(* Logix 5000 project; controller PLC_MCC1300_75F1 vendor 1 type 14 code 166 rev 32.11; software revision 32.04; part 26 of 83 *)
(* tags used below, declared in another part *)
   CM_LineToConveyorStacker_JS2 : CM_LineToConveyorStacker;
   GP_OB_InitializeMain : GP_OB_Initialize;
   M302SpeedUp : MAC_SpeedUp;
   M317 : MAC_Conveyor_Single;
   M317_Data : UDT_Convoy_SL;
   M317_HMW : MAC_Conveyor_HMW;
   M317_M3_ChangeSpeed : BOOL;
   M317_M3_DR_IN_MAJ : MOTION_INSTRUCTION;
   M317_M3_DR_L : AXIS_CIP_DRIVE;
   M317_M3_DR_OUT_MAJ : MOTION_INSTRUCTION;
   M317_M3_DR_OUT_MAS : MOTION_INSTRUCTION;
   M317_M3_DR_OUT_MCD : MOTION_INSTRUCTION;
   M317_SpaceConv_Utilities : SpaceConv_Utilities;
   M350Popup : MAC_Popup_ZC;
   M351 : MAC_Conveyor;
   M351_ALM : MAC_Conveyor_ALM;
   M351_Data : UDT_Convoy_SL;
   M351_HMR : MAC_Conveyor_HMR;
   M351_HMW : MAC_Conveyor_HMW;
   M351_M1_DR : AXIS_CIP_DRIVE;
   M351_M1_DR_IN_MAJ : MOTION_INSTRUCTION;
   M351_M1_DR_IN_MAR : MOTION_INSTRUCTION;
   M351_M1_DR_IN_MAS : MOTION_INSTRUCTION;
   M351_M1_DR_IN_MRP : MOTION_INSTRUCTION;
   M351_M1_DR_MAFR : MOTION_INSTRUCTION;
   M351_M1_DR_MDR : MOTION_INSTRUCTION;
   M351_M1_DR_MSF : MOTION_INSTRUCTION;
   M351_M1_DR_MSO : MOTION_INSTRUCTION;
   M351_M1_DR_OUT_MAJ : MOTION_INSTRUCTION;
   M351_M1_DR_OUT_MAM : MOTION_INSTRUCTION;
   M351_M1_DR_OUT_MAR : MOTION_INSTRUCTION;
   M351_M1_DR_OUT_MAS : MOTION_INSTRUCTION;
   M351_M1_DR_OUT_MCD : MOTION_INSTRUCTION;
   M351_M1_DR_OUT_MRP : MOTION_INSTRUCTION;
   M351_SpaceConv_Utilities : SpaceConv_Utilities;
   M352 : MAC_Conveyor;
   TMP_d : DINT;
   TMP_dDirection : DINT;
   TMP_r : REAL;
   TMP_rAcc : REAL;
   TMP_rDec : REAL;
   TMP_rSpeed : REAL;
   TMP_rTarget_M2 : REAL;
   TMP_xForwardCommadnForCleaningZone : BOOL;
   TMP_xPositioning : BOOL;
   TMP_xPositioning_M2 : BOOL;
   TMP_xPositioning_M3 : BOOL;
   TMP_xPowerSaving : BOOL;
   TMP_xReverse : BOOL;
   TMP_xReverse_M2 : BOOL;
   TMP_xReverse_M3 : BOOL;
   TMP_xRun : BOOL;
   TMP_xRun_M2 : BOOL;
   TMP_xRun_M3 : BOOL;
   xAlwaysOFF : BOOL;
   xDebugOFF : BOOL;
   Z300_Conveyor : UDT_StandConv[29];
   Z300_Conveyor_Conf : UDT_Conveyor_Config[29];
   Z300_Conveyor_HMW : MAC_Conveyor_ZC_HMW[29];
   Z300_Conveyor_IN_MOTION : MAC_Conveyor_ZC_IN_MOTION[29];
   Z301_HMR : MAC_Zone_ML_HMR;
   Z402 : MAC_Zone;
   Z900 : MAC_Zone;
   Z900_HMW : MAC_Zone_HMW;
(* CommandLogic, continued *)

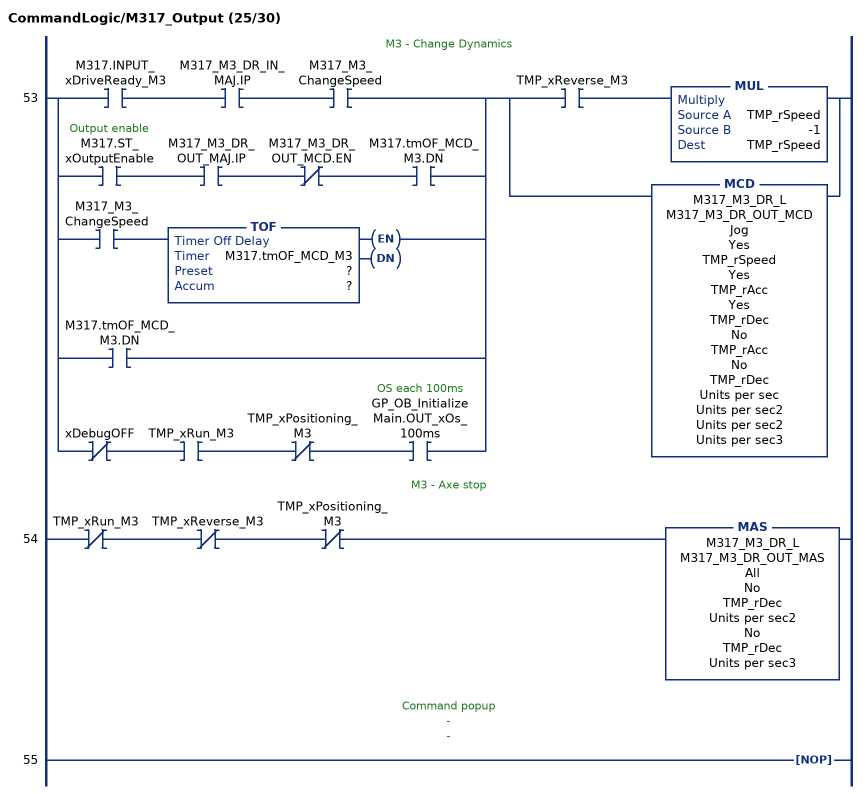
   [picture p307: CommandLogic/M317_Output rungs 53-55]
   // M3 - Change Dynamics
   53: [XIC(M317.INPUT_xDriveReady_M3) XIC(M317_M3_DR_IN_MAJ.IP) XIC(M317_M3_ChangeSpeed) ,XIC(M317.ST_xOutputEnable) XIC(M317_M3_DR_OUT_MAJ.IP) XIO(M317_M3_DR_OUT_MCD.EN) XIC(M317.tmOF_MCD_M3.DN) ,[XIC(M317_M3_ChangeSpeed) TOF(M317.tmOF_MCD_M3,?,?) ,XIC(M317.tmOF_MCD_M3.DN) ] ,XIO(xDebugOFF) XIC(TMP_xRun_M3) XIO(TMP_xPositioning_M3) XIC(GP_OB_InitializeMain.OUT_xOs_100ms) ][XIC(TMP_xReverse_M3) MUL(TMP_rSpeed,-1,TMP_rSpeed) ,MCD(M317_M3_DR_L,M317_M3_DR_OUT_MCD,Jog,Yes,TMP_rSpeed,Yes,TMP_rAcc,Yes,TMP_rDec,No,TMP_rAcc,No,TMP_rDec,Units per sec,Units per sec2,Units per sec2,Units per sec3) ];
   // M3 - Axe stop
   54: XIO(TMP_xRun_M3)XIO(TMP_xReverse_M3)XIO(TMP_xPositioning_M3)MAS(M317_M3_DR_L,M317_M3_DR_OUT_MAS,All,No,TMP_rDec,Units per sec2,No,TMP_rDec,Units per sec3);
   // Command popup
   // -
   // -
   55: NOP();
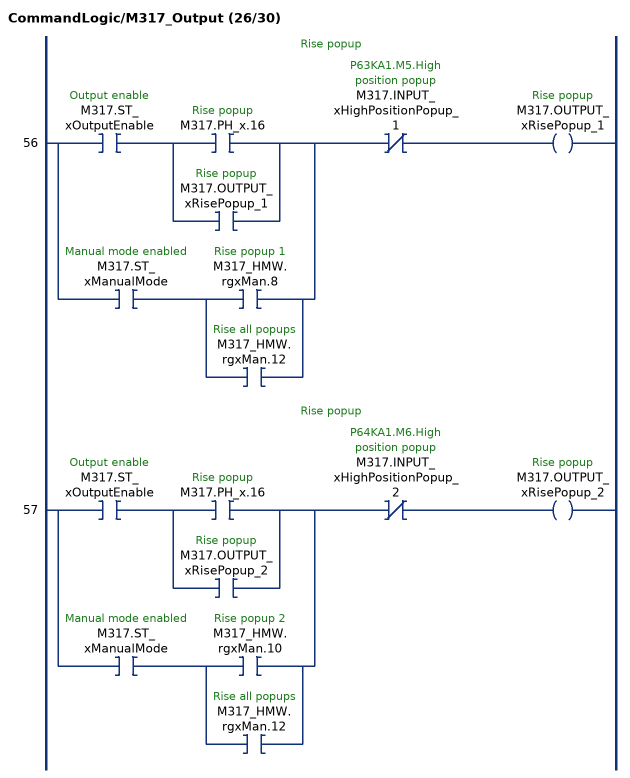
   // Rise popup
   56: [XIC(M317.ST_xOutputEnable) [XIC(M317.PH_x.16) ,XIC(M317.OUTPUT_xRisePopup_1) ] ,XIC(M317.ST_xManualMode) [XIC(M317_HMW.rgxMan.8) ,XIC(M317_HMW.rgxMan.12) ] ]XIO(M317.INPUT_xHighPositionPopup_1)OTE(M317.OUTPUT_xRisePopup_1);
   // Rise popup
   57: [XIC(M317.ST_xOutputEnable) [XIC(M317.PH_x.16) ,XIC(M317.OUTPUT_xRisePopup_2) ] ,XIC(M317.ST_xManualMode) [XIC(M317_HMW.rgxMan.10) ,XIC(M317_HMW.rgxMan.12) ] ]XIO(M317.INPUT_xHighPositionPopup_2)OTE(M317.OUTPUT_xRisePopup_2);
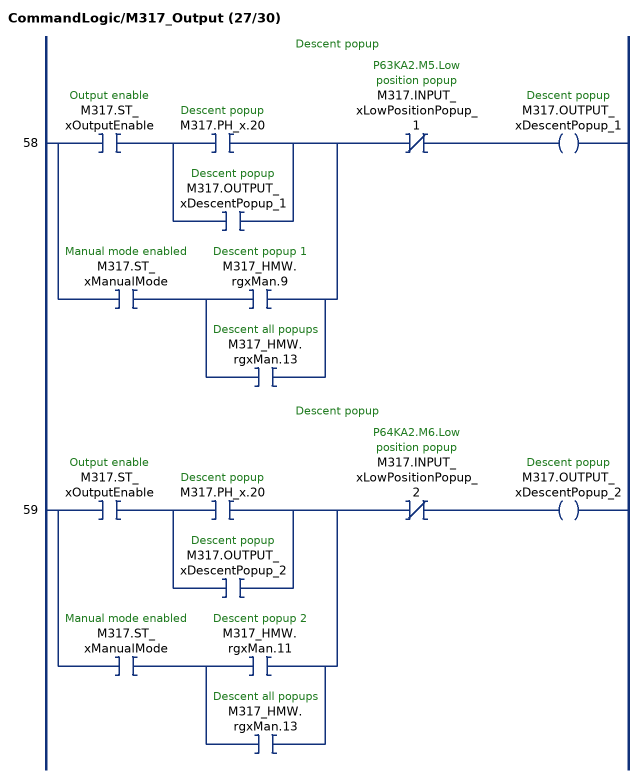
   // Descent popup
   58: [XIC(M317.ST_xOutputEnable) [XIC(M317.PH_x.20) ,XIC(M317.OUTPUT_xDescentPopup_1) ] ,XIC(M317.ST_xManualMode) [XIC(M317_HMW.rgxMan.9) ,XIC(M317_HMW.rgxMan.13) ] ]XIO(M317.INPUT_xLowPositionPopup_1)OTE(M317.OUTPUT_xDescentPopup_1);
   // Descent popup
   59: [XIC(M317.ST_xOutputEnable) [XIC(M317.PH_x.20) ,XIC(M317.OUTPUT_xDescentPopup_2) ] ,XIC(M317.ST_xManualMode) [XIC(M317_HMW.rgxMan.11) ,XIC(M317_HMW.rgxMan.13) ] ]XIO(M317.INPUT_xLowPositionPopup_2)OTE(M317.OUTPUT_xDescentPopup_2);
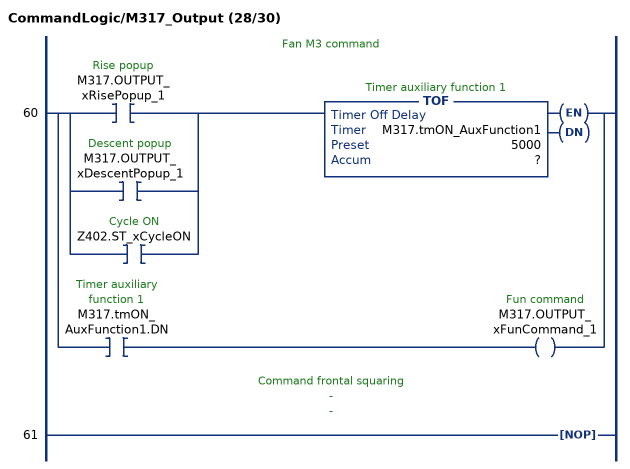
   // Fan M3 command
   60: [[XIC(M317.OUTPUT_xRisePopup_1) ,[XIC(M317.OUTPUT_xDescentPopup_1) ,XIC(Z402.ST_xCycleON) ] ] TOF(M317.tmON_AuxFunction1,?,?) ,XIC(M317.tmON_AuxFunction1.DN) OTE(M317.OUTPUT_xFunCommand_1) ];
   // Command frontal squaring
   // -
   // -
   61: NOP();
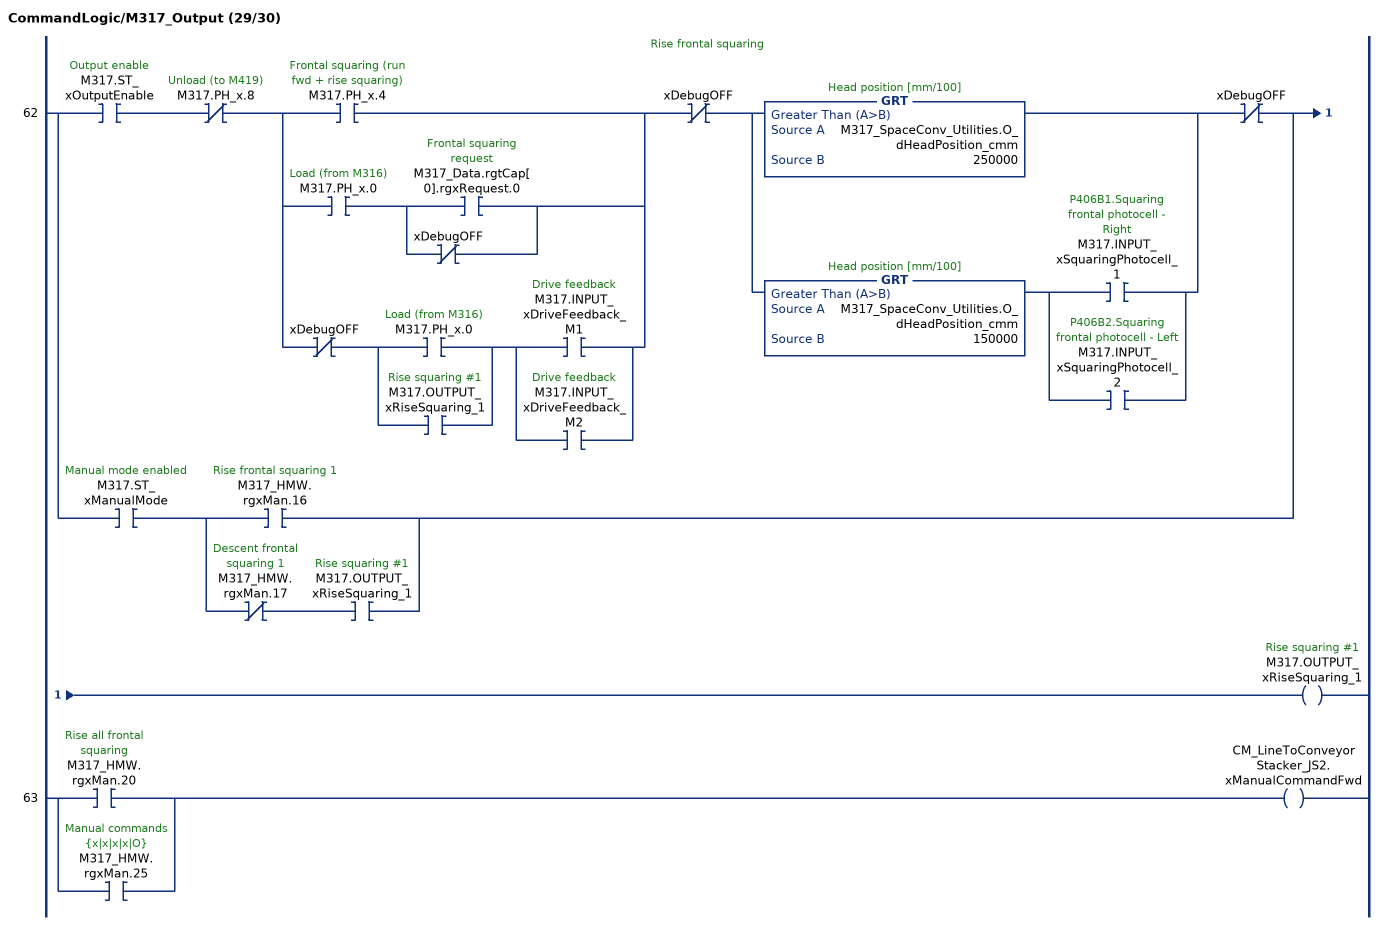
   // Rise frontal squaring
   62: [XIC(M317.ST_xOutputEnable) XIO(M317.PH_x.8) [XIC(M317.PH_x.4) ,XIC(M317.PH_x.0) [XIC(M317_Data.rgtCap[0].rgxRequest.0) ,XIO(xDebugOFF) ] ,XIO(xDebugOFF) [XIC(M317.PH_x.0) ,XIC(M317.OUTPUT_xRiseSquaring_1) ] [XIC(M317.INPUT_xDriveFeedback_M1) ,XIC(M317.INPUT_xDriveFeedback_M2) ] ] XIO(xDebugOFF) [GRT(M317_SpaceConv_Utilities.O_dHeadPosition_cmm,250000) ,GRT(M317_SpaceConv_Utilities.O_dHeadPosition_cmm,150000) [XIC(M317.INPUT_xSquaringPhotocell_1) ,XIC(M317.INPUT_xSquaringPhotocell_2) ] ] XIO(xDebugOFF) ,XIC(M317.ST_xManualMode) [XIC(M317_HMW.rgxMan.16) ,XIO(M317_HMW.rgxMan.17) XIC(M317.OUTPUT_xRiseSquaring_1) ] ]OTE(M317.OUTPUT_xRiseSquaring_1);
   63: [XIC(M317_HMW.rgxMan.20) ,XIC(M317_HMW.rgxMan.25) ]OTE(CM_LineToConveyorStacker_JS2.xManualCommandFwd);
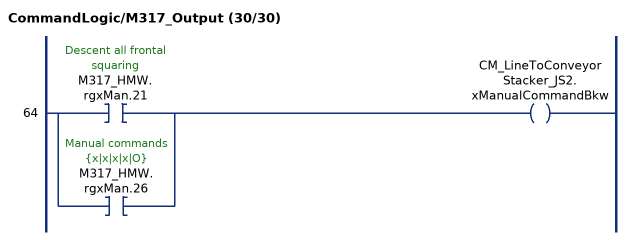
   64: [XIC(M317_HMW.rgxMan.21) ,XIC(M317_HMW.rgxMan.26) ]OTE(CM_LineToConveyorStacker_JS2.xManualCommandBkw);
END_ROUTINE

ROUTINE M350M1_Conveyor_Output   (* ladder *)
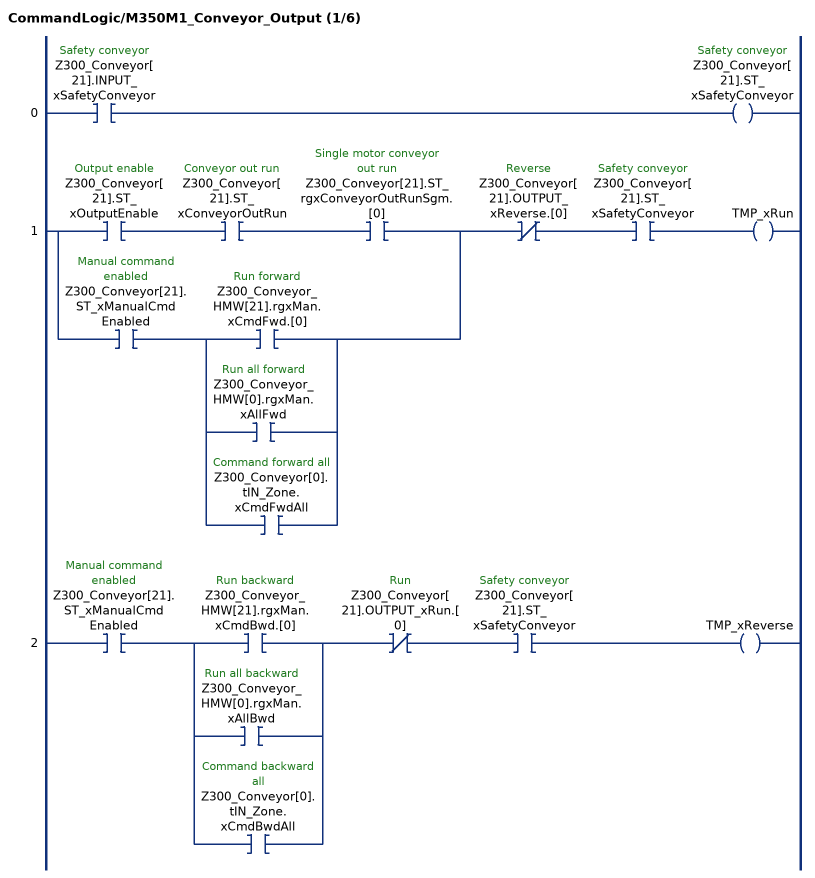
   0: XIC(Z300_Conveyor[21].INPUT_xSafetyConveyor)OTE(Z300_Conveyor[21].ST_xSafetyConveyor);
   1: [XIC(Z300_Conveyor[21].ST_xOutputEnable) XIC(Z300_Conveyor[21].ST_xConveyorOutRun) XIC(Z300_Conveyor[21].ST_rgxConveyorOutRunSgm.[0]) ,XIC(Z300_Conveyor[21].ST_xManualCmdEnabled) [XIC(Z300_Conveyor_HMW[21].rgxMan.xCmdFwd.[0]) ,XIC(Z300_Conveyor_HMW[0].rgxMan.xAllFwd) ,XIC(Z300_Conveyor[0].tIN_Zone.xCmdFwdAll) ] ]XIO(Z300_Conveyor[21].OUTPUT_xReverse.[0])XIC(Z300_Conveyor[21].ST_xSafetyConveyor)OTE(TMP_xRun);
   2: XIC(Z300_Conveyor[21].ST_xManualCmdEnabled)[XIC(Z300_Conveyor_HMW[21].rgxMan.xCmdBwd.[0]) ,XIC(Z300_Conveyor_HMW[0].rgxMan.xAllBwd) ,XIC(Z300_Conveyor[0].tIN_Zone.xCmdBwdAll) ]XIO(Z300_Conveyor[21].OUTPUT_xRun.[0])XIC(Z300_Conveyor[21].ST_xSafetyConveyor)OTE(TMP_xReverse);
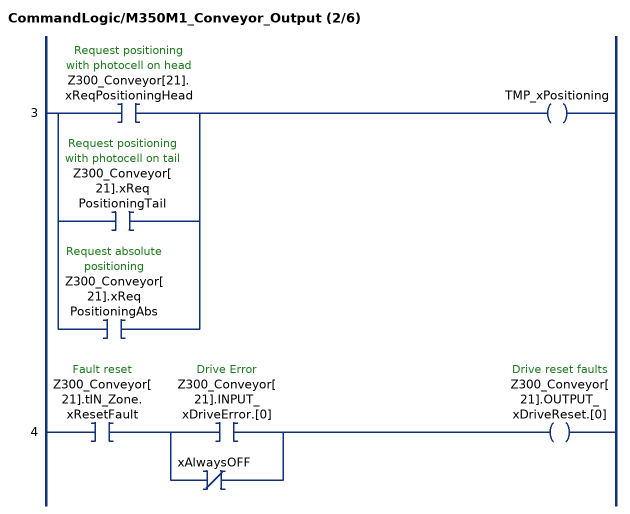
   3: [XIC(Z300_Conveyor[21].xReqPositioningHead) ,XIC(Z300_Conveyor[21].xReqPositioningTail) ,XIC(Z300_Conveyor[21].xReqPositioningAbs) ]OTE(TMP_xPositioning);
   4: XIC(Z300_Conveyor[21].tIN_Zone.xResetFault)[XIC(Z300_Conveyor[21].INPUT_xDriveError.[0]) ,XIO(xAlwaysOFF) ]OTE(Z300_Conveyor[21].OUTPUT_xDriveReset.[0]);
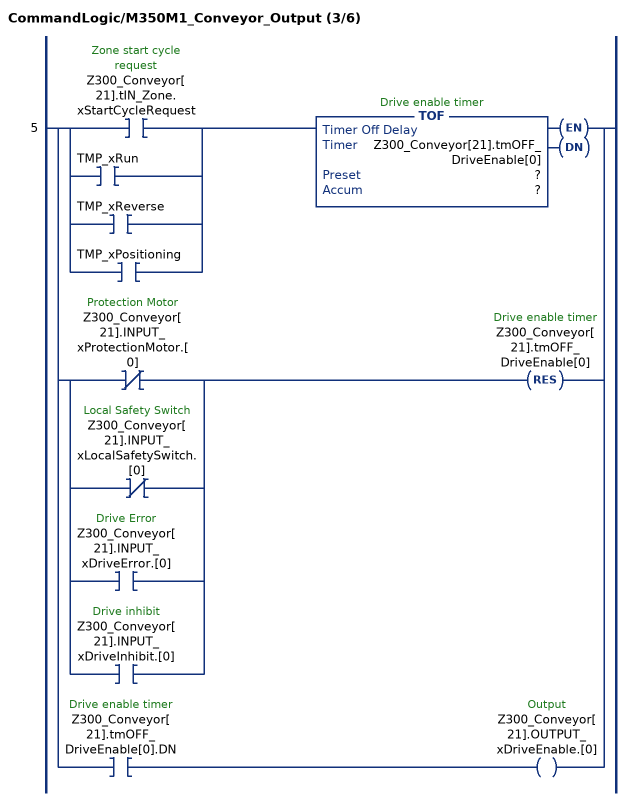
   5: [[XIC(Z300_Conveyor[21].tIN_Zone.xStartCycleRequest) ,XIC(TMP_xRun) ,XIC(TMP_xReverse) ,XIC(TMP_xPositioning) ] TOF(Z300_Conveyor[21].tmOFF_DriveEnable[0],?,?) ,[XIO(Z300_Conveyor[21].INPUT_xProtectionMotor.[0]) ,XIO(Z300_Conveyor[21].INPUT_xLocalSafetySwitch.[0]) ,XIC(Z300_Conveyor[21].INPUT_xDriveError.[0]) ,XIC(Z300_Conveyor[21].INPUT_xDriveInhibit.[0]) ] RES(Z300_Conveyor[21].tmOFF_DriveEnable[0]) ,XIC(Z300_Conveyor[21].tmOFF_DriveEnable[0].DN) OTE(Z300_Conveyor[21].OUTPUT_xDriveEnable.[0]) ];
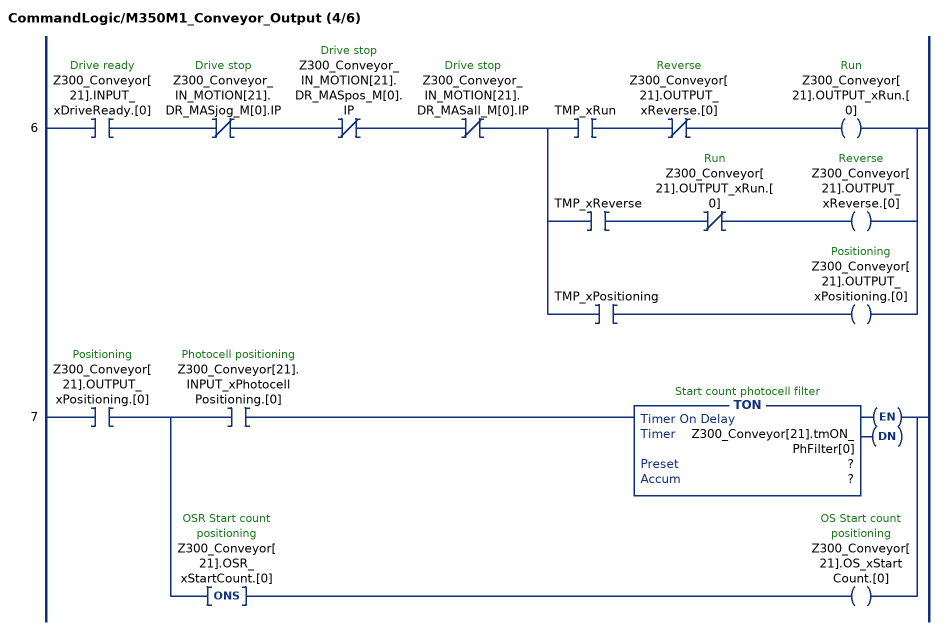
   6: XIC(Z300_Conveyor[21].INPUT_xDriveReady.[0])XIO(Z300_Conveyor_IN_MOTION[21].DR_MASjog_M[0].IP)XIO(Z300_Conveyor_IN_MOTION[21].DR_MASpos_M[0].IP)XIO(Z300_Conveyor_IN_MOTION[21].DR_MASall_M[0].IP)[XIC(TMP_xRun) XIO(Z300_Conveyor[21].OUTPUT_xReverse.[0]) OTE(Z300_Conveyor[21].OUTPUT_xRun.[0]) ,XIC(TMP_xReverse) XIO(Z300_Conveyor[21].OUTPUT_xRun.[0]) OTE(Z300_Conveyor[21].OUTPUT_xReverse.[0]) ,XIC(TMP_xPositioning) OTE(Z300_Conveyor[21].OUTPUT_xPositioning.[0]) ];
   7: XIC(Z300_Conveyor[21].OUTPUT_xPositioning.[0])[XIC(Z300_Conveyor[21].INPUT_xPhotocellPositioning.[0]) TON(Z300_Conveyor[21].tmON_PhFilter[0],?,?) ,ONS(Z300_Conveyor[21].OSR_xStartCount.[0]) OTE(Z300_Conveyor[21].OS_xStartCount.[0]) ];
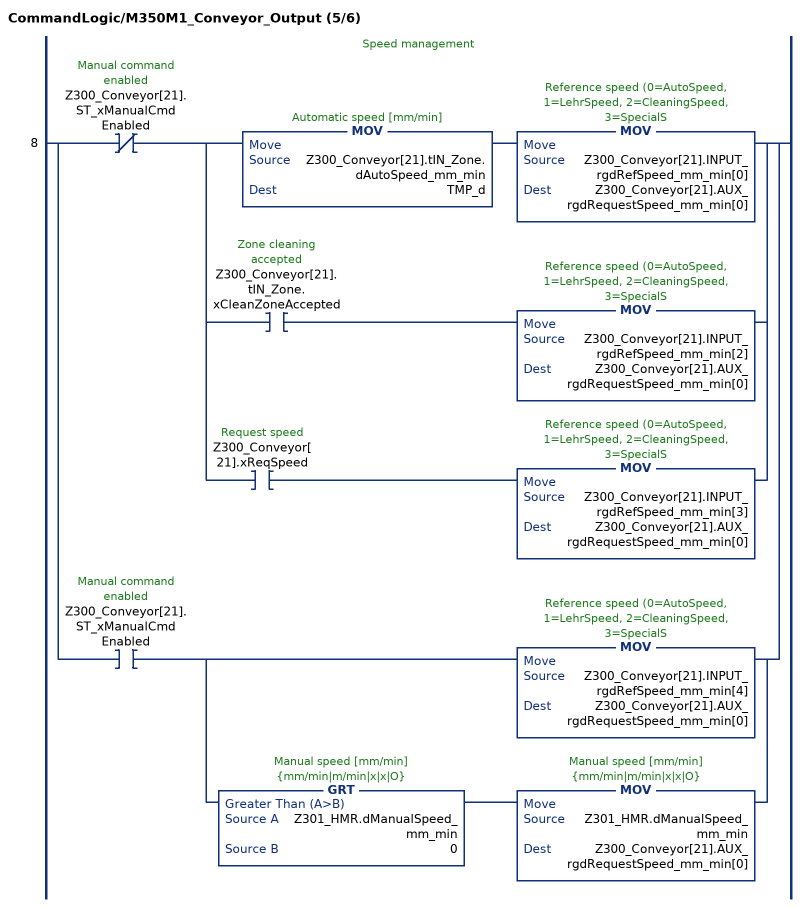
   // Speed management
   8: [XIO(Z300_Conveyor[21].ST_xManualCmdEnabled) [MOV(Z300_Conveyor[21].tIN_Zone.dAutoSpeed_mm_min,TMP_d) MOV(Z300_Conveyor[21].INPUT_rgdRefSpeed_mm_min[0],Z300_Conveyor[21].AUX_rgdRequestSpeed_mm_min[0]) ,XIC(Z300_Conveyor[21].tIN_Zone.xCleanZoneAccepted) MOV(Z300_Conveyor[21].INPUT_rgdRefSpeed_mm_min[2],Z300_Conveyor[21].AUX_rgdRequestSpeed_mm_min[0]) ,XIC(Z300_Conveyor[21].xReqSpeed) MOV(Z300_Conveyor[21].INPUT_rgdRefSpeed_mm_min[3],Z300_Conveyor[21].AUX_rgdRequestSpeed_mm_min[0]) ] ,XIC(Z300_Conveyor[21].ST_xManualCmdEnabled) [MOV(Z300_Conveyor[21].INPUT_rgdRefSpeed_mm_min[4],Z300_Conveyor[21].AUX_rgdRequestSpeed_mm_min[0]) ,GRT(Z301_HMR.dManualSpeed_mm_min,0) MOV(Z301_HMR.dManualSpeed_mm_min,Z300_Conveyor[21].AUX_rgdRequestSpeed_mm_min[0]) ] ];
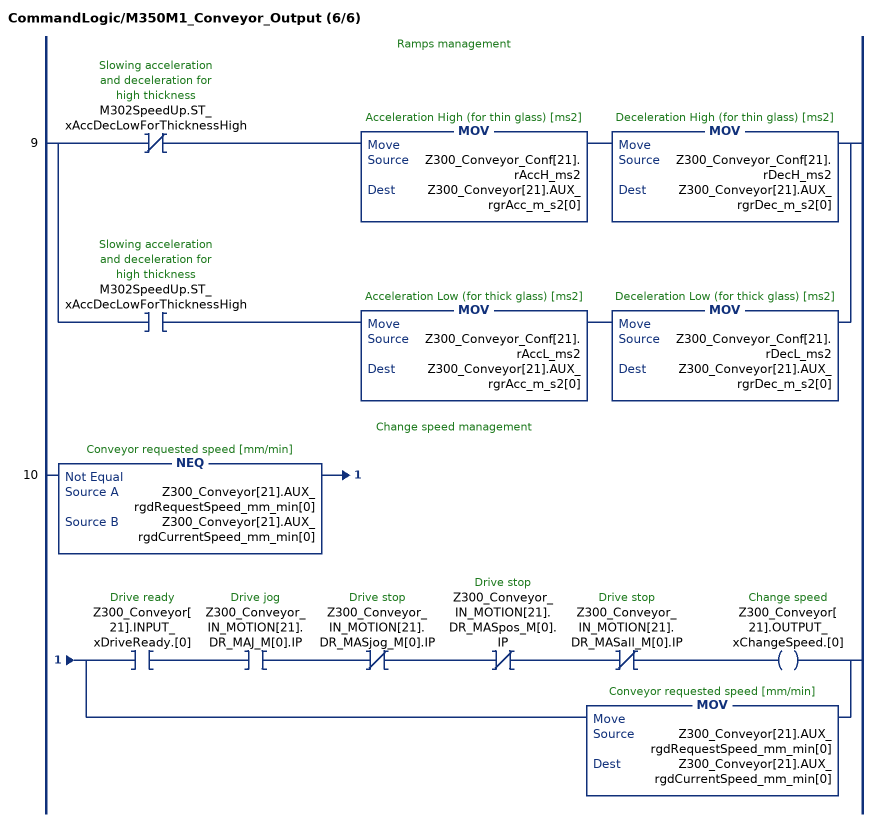
   // Ramps management
   9: [XIO(M302SpeedUp.ST_xAccDecLowForThicknessHigh) MOV(Z300_Conveyor_Conf[21].rAccH_ms2,Z300_Conveyor[21].AUX_rgrAcc_m_s2[0]) MOV(Z300_Conveyor_Conf[21].rDecH_ms2,Z300_Conveyor[21].AUX_rgrDec_m_s2[0]) ,XIC(M302SpeedUp.ST_xAccDecLowForThicknessHigh) MOV(Z300_Conveyor_Conf[21].rAccL_ms2,Z300_Conveyor[21].AUX_rgrAcc_m_s2[0]) MOV(Z300_Conveyor_Conf[21].rDecL_ms2,Z300_Conveyor[21].AUX_rgrDec_m_s2[0]) ];
   // Change speed management
   10: NEQ(Z300_Conveyor[21].AUX_rgdRequestSpeed_mm_min[0],Z300_Conveyor[21].AUX_rgdCurrentSpeed_mm_min[0])[XIC(Z300_Conveyor[21].INPUT_xDriveReady.[0]) XIC(Z300_Conveyor_IN_MOTION[21].DR_MAJ_M[0].IP) XIO(Z300_Conveyor_IN_MOTION[21].DR_MASjog_M[0].IP) XIO(Z300_Conveyor_IN_MOTION[21].DR_MASpos_M[0].IP) XIO(Z300_Conveyor_IN_MOTION[21].DR_MASall_M[0].IP) OTE(Z300_Conveyor[21].OUTPUT_xChangeSpeed.[0]) ,MOV(Z300_Conveyor[21].AUX_rgdRequestSpeed_mm_min[0],Z300_Conveyor[21].AUX_rgdCurrentSpeed_mm_min[0]) ];
END_ROUTINE

ROUTINE M351_Output   (* ladder *)
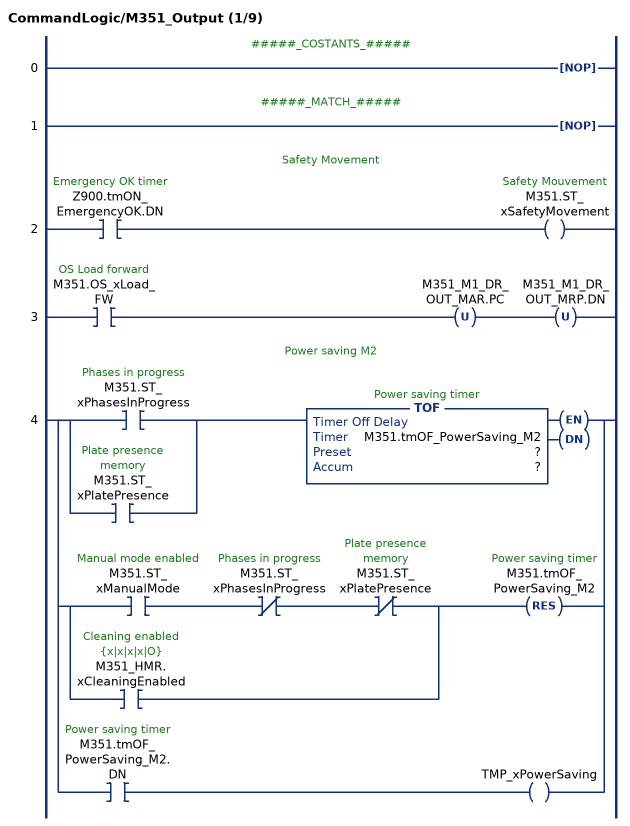
   // #####_COSTANTS_#####
   0: NOP();
   // #####_MATCH_#####
   1: NOP();
   // Safety Movement
   2: XIC(Z900.tmON_EmergencyOK.DN)OTE(M351.ST_xSafetyMovement);
   3: XIC(M351.OS_xLoad_FW)OTU(M351_M1_DR_OUT_MAR.PC)OTU(M351_M1_DR_OUT_MRP.DN);
   // Power saving M2
   4: [[XIC(M351.ST_xPhasesInProgress) ,XIC(M351.ST_xPlatePresence) ] TOF(M351.tmOF_PowerSaving_M2,?,?) ,[XIC(M351.ST_xManualMode) XIO(M351.ST_xPhasesInProgress) XIO(M351.ST_xPlatePresence) ,XIC(M351_HMR.xCleaningEnabled) ] RES(M351.tmOF_PowerSaving_M2) ,XIC(M351.tmOF_PowerSaving_M2.DN) OTE(TMP_xPowerSaving) ];
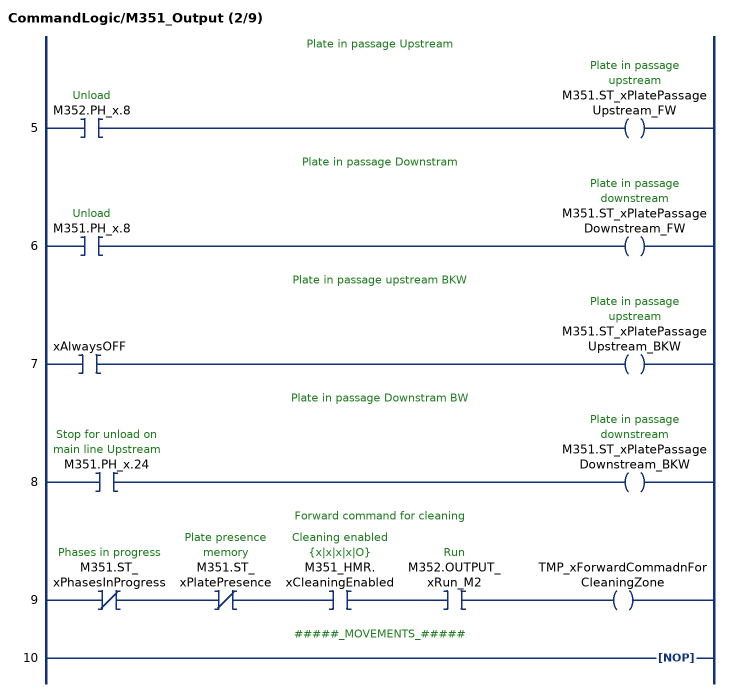
   // Plate in passage Upstream
   5: XIC(M352.PH_x.8)OTE(M351.ST_xPlatePassageUpstream_FW);
   // Plate in passage Downstram
   6: XIC(M351.PH_x.8)OTE(M351.ST_xPlatePassageDownstream_FW);
   // Plate in passage upstream BKW
   7: XIC(xAlwaysOFF)OTE(M351.ST_xPlatePassageUpstream_BKW);
   // Plate in passage Downstram BW
   8: XIC(M351.PH_x.24)OTE(M351.ST_xPlatePassageDownstream_BKW);
   // Forward command for cleaning
   9: XIO(M351.ST_xPhasesInProgress)XIO(M351.ST_xPlatePresence)XIC(M351_HMR.xCleaningEnabled)XIC(M352.OUTPUT_xRun_M2)OTE(TMP_xForwardCommadnForCleaningZone);
   // #####_MOVEMENTS_#####
   10: NOP();
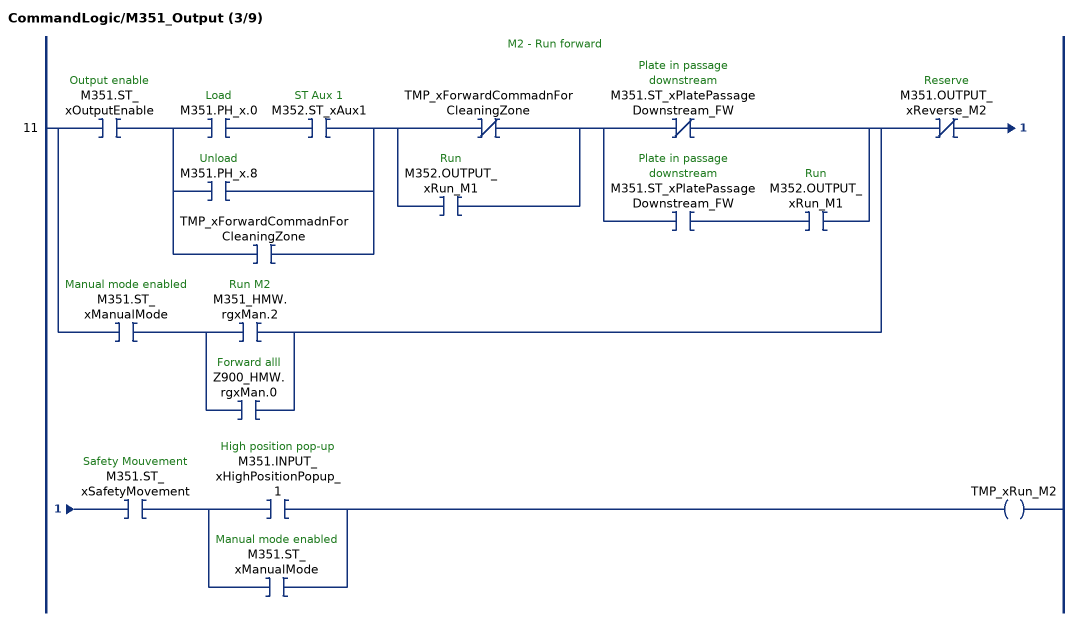
   // M2 - Run forward
   11: [XIC(M351.ST_xOutputEnable) [XIC(M351.PH_x.0) XIC(M352.ST_xAux1) ,XIC(M351.PH_x.8) ,XIC(TMP_xForwardCommadnForCleaningZone) ] [XIO(TMP_xForwardCommadnForCleaningZone) ,XIC(M352.OUTPUT_xRun_M1) ] [XIO(M351.ST_xPlatePassageDownstream_FW) ,XIC(M351.ST_xPlatePassageDownstream_FW) XIC(M352.OUTPUT_xRun_M1) ] ,XIC(M351.ST_xManualMode) [XIC(M351_HMW.rgxMan.2) ,XIC(Z900_HMW.rgxMan.0) ] ]XIO(M351.OUTPUT_xReverse_M2)XIC(M351.ST_xSafetyMovement)[XIC(M351.INPUT_xHighPositionPopup_1) ,XIC(M351.ST_xManualMode) ]OTE(TMP_xRun_M2);
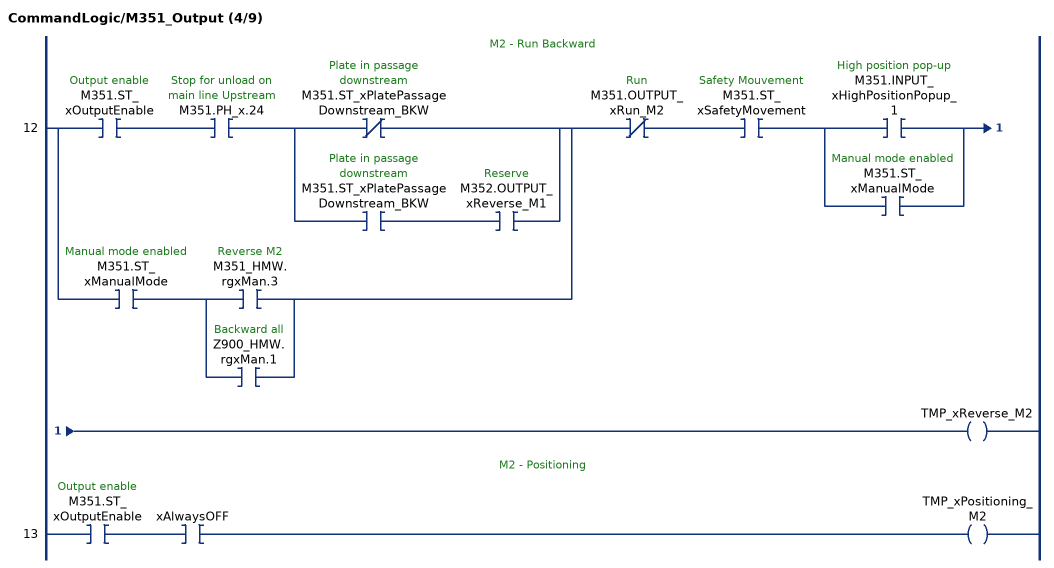
   // M2 - Run Backward
   12: [XIC(M351.ST_xOutputEnable) XIC(M351.PH_x.24) [XIO(M351.ST_xPlatePassageDownstream_BKW) ,XIC(M351.ST_xPlatePassageDownstream_BKW) XIC(M352.OUTPUT_xReverse_M1) ] ,XIC(M351.ST_xManualMode) [XIC(M351_HMW.rgxMan.3) ,XIC(Z900_HMW.rgxMan.1) ] ]XIO(M351.OUTPUT_xRun_M2)XIC(M351.ST_xSafetyMovement)[XIC(M351.INPUT_xHighPositionPopup_1) ,XIC(M351.ST_xManualMode) ]OTE(TMP_xReverse_M2);
   // M2 - Positioning
   13: XIC(M351.ST_xOutputEnable)XIC(xAlwaysOFF)OTE(TMP_xPositioning_M2);
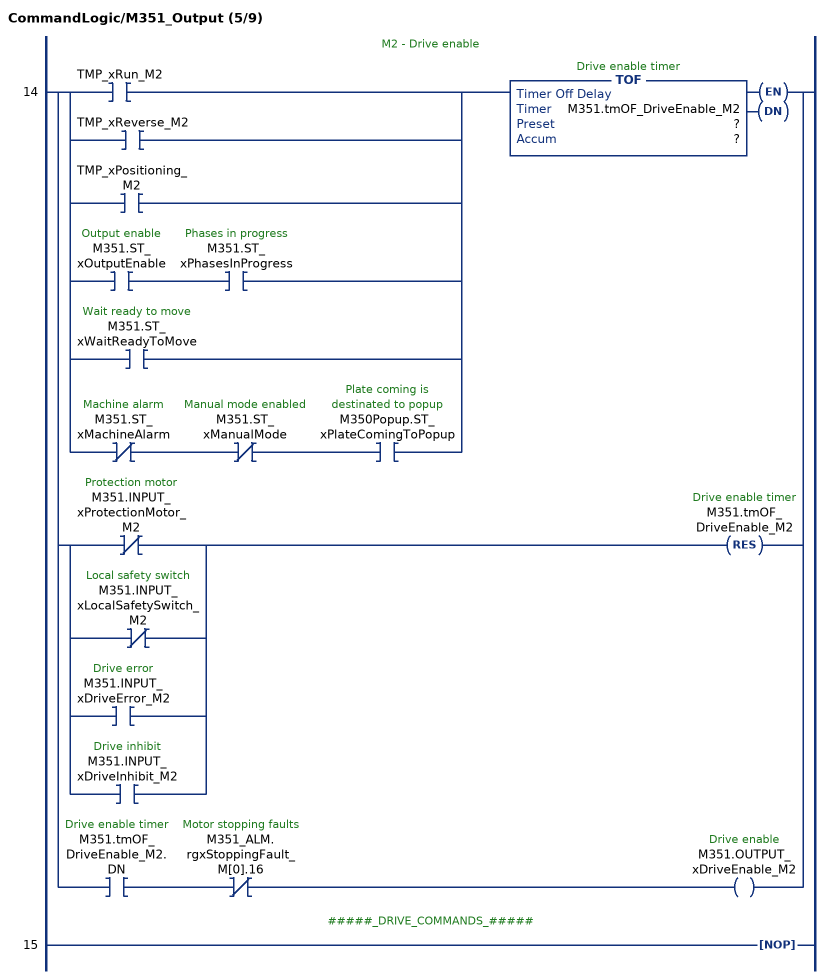
   // M2 - Drive enable
   14: [[XIC(TMP_xRun_M2) ,XIC(TMP_xReverse_M2) ,XIC(TMP_xPositioning_M2) ,XIC(M351.ST_xOutputEnable) XIC(M351.ST_xPhasesInProgress) ,XIC(M351.ST_xWaitReadyToMove) ,XIO(M351.ST_xMachineAlarm) XIO(M351.ST_xManualMode) XIC(M350Popup.ST_xPlateComingToPopup) ] TOF(M351.tmOF_DriveEnable_M2,?,?) ,[XIO(M351.INPUT_xProtectionMotor_M2) ,XIO(M351.INPUT_xLocalSafetySwitch_M2) ,XIC(M351.INPUT_xDriveError_M2) ,XIC(M351.INPUT_xDriveInhibit_M2) ] RES(M351.tmOF_DriveEnable_M2) ,XIC(M351.tmOF_DriveEnable_M2.DN) XIO(M351_ALM.rgxStoppingFault_M[0].16) OTE(M351.OUTPUT_xDriveEnable_M2) ];
   // #####_DRIVE_COMMANDS_#####
   15: NOP();
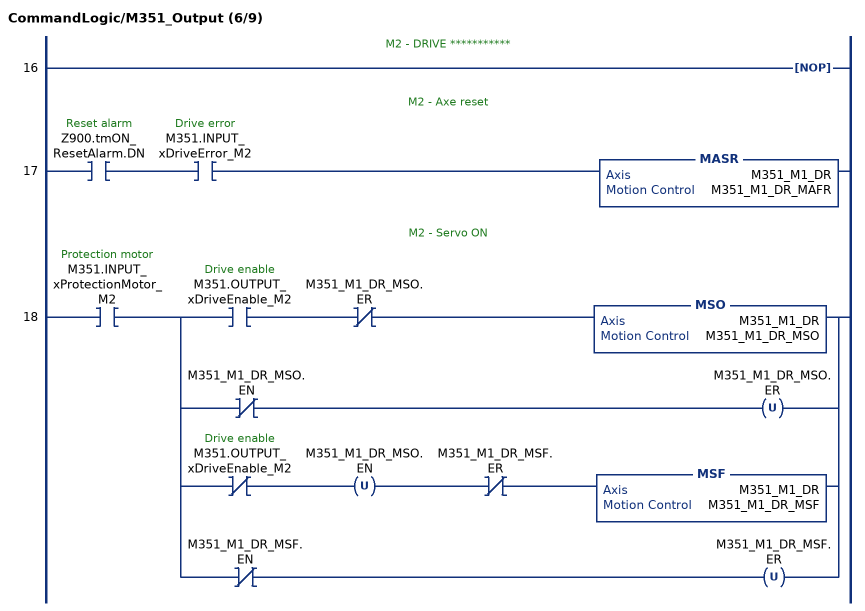
   // M2 - DRIVE ***********
   16: NOP();
   // M2 - Axe reset
   17: XIC(Z900.tmON_ResetAlarm.DN)XIC(M351.INPUT_xDriveError_M2)MASR(M351_M1_DR,M351_M1_DR_MAFR);
   // M2 - Servo ON
   18: XIC(M351.INPUT_xProtectionMotor_M2)[XIC(M351.OUTPUT_xDriveEnable_M2) XIO(M351_M1_DR_MSO.ER) MSO(M351_M1_DR,M351_M1_DR_MSO) ,XIO(M351_M1_DR_MSO.EN) OTU(M351_M1_DR_MSO.ER) ,XIO(M351.OUTPUT_xDriveEnable_M2) OTU(M351_M1_DR_MSO.EN) XIO(M351_M1_DR_MSF.ER) MSF(M351_M1_DR,M351_M1_DR_MSF) ,XIO(M351_M1_DR_MSF.EN) OTU(M351_M1_DR_MSF.ER) ];
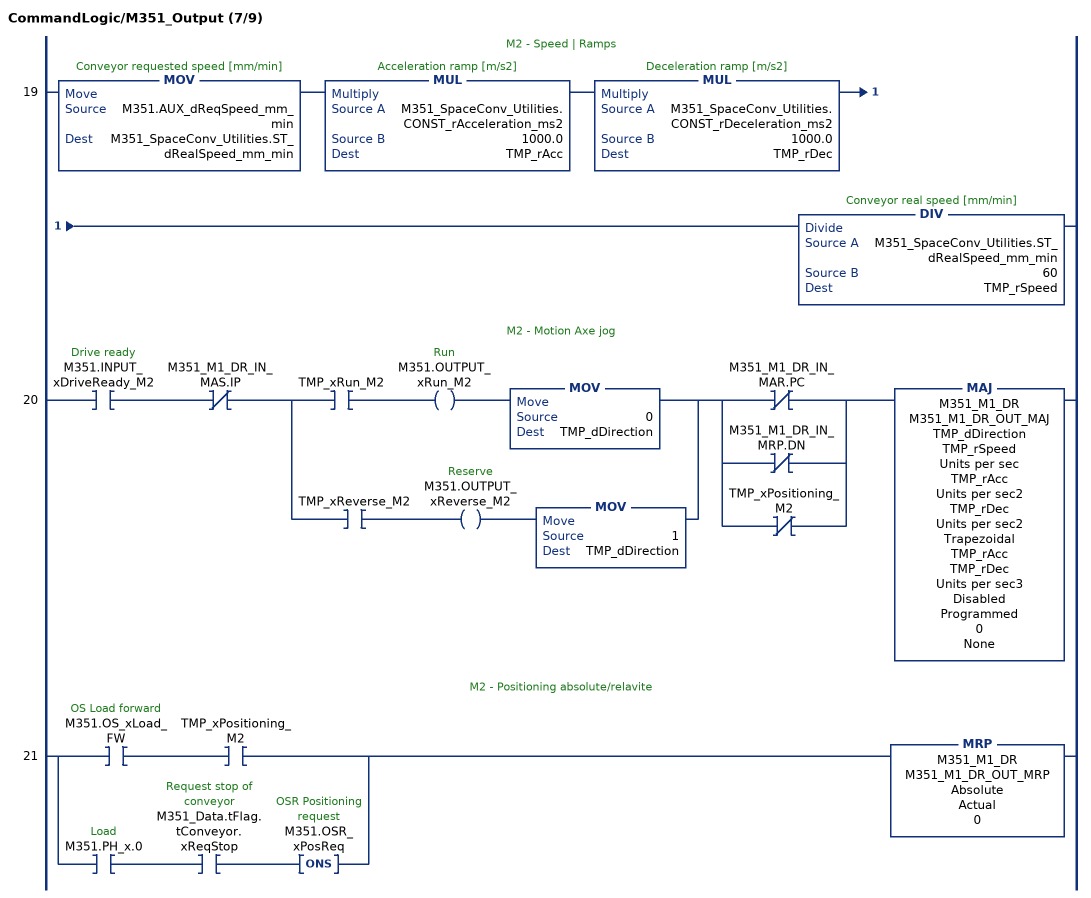
   // M2 - Speed | Ramps
   19: MOV(M351.AUX_dReqSpeed_mm_min,M351_SpaceConv_Utilities.ST_dRealSpeed_mm_min)MUL(M351_SpaceConv_Utilities.CONST_rAcceleration_ms2,1000.0,TMP_rAcc)MUL(M351_SpaceConv_Utilities.CONST_rDeceleration_ms2,1000.0,TMP_rDec)DIV(M351_SpaceConv_Utilities.ST_dRealSpeed_mm_min,60,TMP_rSpeed);
   // M2 - Motion Axe jog
   20: XIC(M351.INPUT_xDriveReady_M2)XIO(M351_M1_DR_IN_MAS.IP)[XIC(TMP_xRun_M2) OTE(M351.OUTPUT_xRun_M2) MOV(0,TMP_dDirection) ,XIC(TMP_xReverse_M2) OTE(M351.OUTPUT_xReverse_M2) MOV(1,TMP_dDirection) ][XIO(M351_M1_DR_IN_MAR.PC) ,XIO(M351_M1_DR_IN_MRP.DN) ,XIO(TMP_xPositioning_M2) ]MAJ(M351_M1_DR,M351_M1_DR_OUT_MAJ,TMP_dDirection,TMP_rSpeed,Units per sec,TMP_rAcc,Units per sec2,TMP_rDec,Units per sec2,Trapezoidal,TMP_rAcc,TMP_rDec,Units per sec3,Disabled,Programmed,0,None);
   // M2 - Positioning absolute/relavite
   21: [XIC(M351.OS_xLoad_FW) XIC(TMP_xPositioning_M2) ,XIC(M351.PH_x.0) XIC(M351_Data.tFlag.tConveyor.xReqStop) ONS(M351.OSR_xPosReq) ]MRP(M351_M1_DR,M351_M1_DR_OUT_MRP,Absolute,Actual,0);
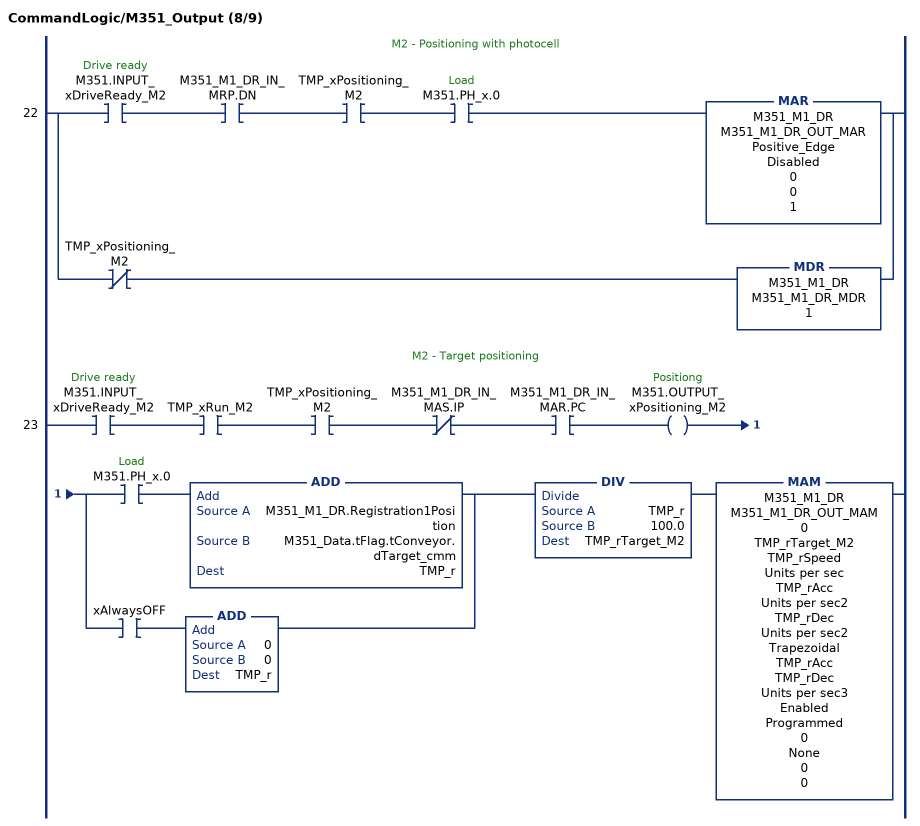
   // M2 - Positioning with photocell
   22: [XIC(M351.INPUT_xDriveReady_M2) XIC(M351_M1_DR_IN_MRP.DN) XIC(TMP_xPositioning_M2) XIC(M351.PH_x.0) MAR(M351_M1_DR,M351_M1_DR_OUT_MAR,Positive_Edge,Disabled,0,0,1) ,XIO(TMP_xPositioning_M2) MDR(M351_M1_DR,M351_M1_DR_MDR,1) ];
   // M2 - Target positioning
   23: XIC(M351.INPUT_xDriveReady_M2)XIC(TMP_xRun_M2)XIC(TMP_xPositioning_M2)XIO(M351_M1_DR_IN_MAS.IP)XIC(M351_M1_DR_IN_MAR.PC)OTE(M351.OUTPUT_xPositioning_M2)[XIC(M351.PH_x.0) ADD(M351_M1_DR.Registration1Position,M351_Data.tFlag.tConveyor.dTarget_cmm,TMP_r) ,XIC(xAlwaysOFF) ADD(0,0,TMP_r) ]DIV(TMP_r,100.0,TMP_rTarget_M2)MAM(M351_M1_DR,M351_M1_DR_OUT_MAM,0,TMP_rTarget_M2,TMP_rSpeed,Units per sec,TMP_rAcc,Units per sec2,TMP_rDec,Units per sec2,Trapezoidal,TMP_rAcc,TMP_rDec,Units per sec3,Enabled,Programmed,0,None,0,0);
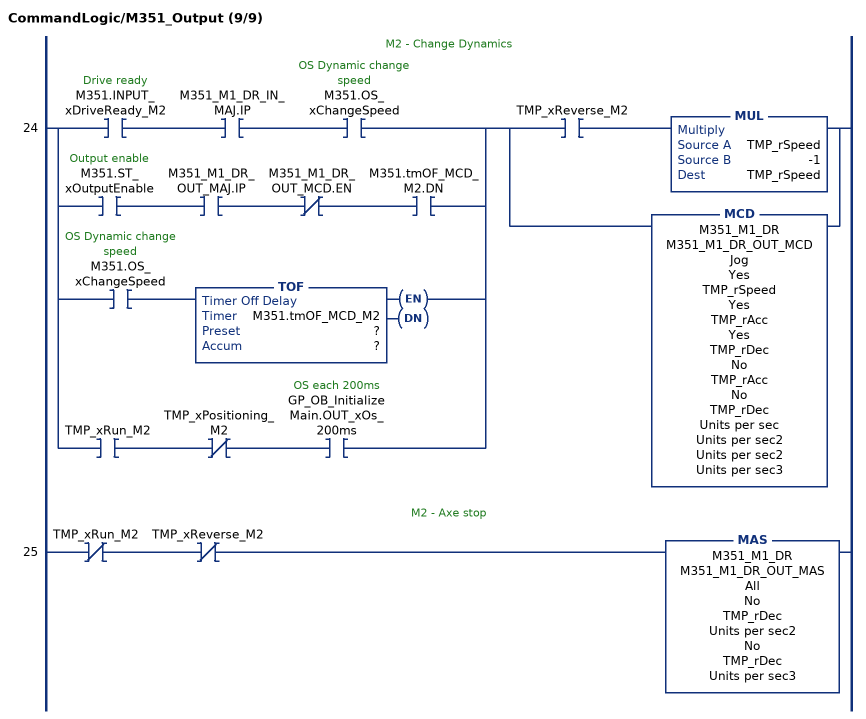
   // M2 - Change Dynamics
   24: [XIC(M351.INPUT_xDriveReady_M2) XIC(M351_M1_DR_IN_MAJ.IP) XIC(M351.OS_xChangeSpeed) ,XIC(M351.ST_xOutputEnable) XIC(M351_M1_DR_OUT_MAJ.IP) XIO(M351_M1_DR_OUT_MCD.EN) XIC(M351.tmOF_MCD_M2.DN) ,XIC(M351.OS_xChangeSpeed) TOF(M351.tmOF_MCD_M2,?,?) ,XIC(TMP_xRun_M2) XIO(TMP_xPositioning_M2) XIC(GP_OB_InitializeMain.OUT_xOs_200ms) ][XIC(TMP_xReverse_M2) MUL(TMP_rSpeed,-1,TMP_rSpeed) ,MCD(M351_M1_DR,M351_M1_DR_OUT_MCD,Jog,Yes,TMP_rSpeed,Yes,TMP_rAcc,Yes,TMP_rDec,No,TMP_rAcc,No,TMP_rDec,Units per sec,Units per sec2,Units per sec2,Units per sec3) ];
   // M2 - Axe stop
   25: XIO(TMP_xRun_M2)XIO(TMP_xReverse_M2)MAS(M351_M1_DR,M351_M1_DR_OUT_MAS,All,No,TMP_rDec,Units per sec2,No,TMP_rDec,Units per sec3);
END_ROUTINE
